VERSION : 0.1
   STRUCT
      SDC_Interlocks_In : "UDT_AB_Interlocks_SDC_In";
      SDC_Interlocks_Out : "UDT_AB_Interlocks_SDC_Out";
      Carrier : Array[1..99] of "UDT_AB_Interlocks_Carrier";
   END_STRUCT;
END_TYPE

TYPE "UDT_AB_Interlocks_SDC_Out"
VERSION : 0.1
   STRUCT
      SDC_Faulted : Bool;
      SDC_Status_1 : Bool;
      SDC_Status_2 : Bool;
      SDC_Status_3 : Bool;
      SDC_Status_4 : Bool;
      SDC_Status_5 : Bool;
      SDC_Status_6 : Bool;
      SDC_Status_7 : Bool;
      SDC_Status_8 : Bool;
      SDC_Status_9 : Bool;
      SDC_Status_10 : Bool;
      SDC_Status_11 : Bool;
      SDC_Status_12 : Bool;
      SDC_Status_13 : Bool;
      SDC_Status_14 : Bool;
      Heartbeat : Bool;
   END_STRUCT;
END_TYPE

// folder: UserDiag

TYPE "UserDiag_typeDevice"
TITLE = UserDiag_typeDevice
VERSION : 0.1
   STRUCT
      hardwareId : Hw_Device := 16#0000;   // Hardware identifier of the device/slave
      number : UInt := 0;   // Profinet device number/Profibus address of the slave
      "name" : String[50];   // Name of the device/slave
      ipAddress : IP_V4;   // IP address of the device
      state : USInt := 0;   // Status of the device/slave. 1:ok; 2:faulty, 3:lost connection, 4:disabled, 5:problem, 12:was faulty, 13:was lost, 14:was disabled, 15:problem gone
      exists : Bool := FALSE;   // TRUE: Device/slave is existing
      configured : Bool := FALSE;   // TRUE: Device/slave is configured
      faulty : Bool := FALSE;   // TRUE: Device/slave is faulty
      problem : Bool := FALSE;   // TRUE: Device/slave has a problem
      disabled : Bool := FALSE;   // TRUE: Device/slave is disabled
      error : Bool := FALSE;   // TRUE: Error in device/slave
      nextDevice : Int;   // device number of next device
      actualConfiguredSlots : Int := 0;   // Number of configured slots in the device/slave
      slots : Array[0.."USERDIAG_SLOTS_PER_DEVICE_UPPER_LIM"] of "UserDiag_typeSlot";   // Slot information of a device/slave
   END_STRUCT;
END_TYPE

TYPE "UserDiag_typeIOSystem"
TITLE = UserDiag_typeIOSystem
VERSION : 0.1
   STRUCT
      hardwareId : Hw_IoSystem := 16#0000;   // Hardware identifier of the IO-System/DP-Mastersystem
      number : UInt := 0;   // IO-System/DP-Mastersystem number
      error : Bool := FALSE;   // TRUE: Error in IO-System/DP-Mastersystem
      firstDevice : Int := 0;   // device number (index) of first device in IO System
      lastDevice : Int := 0;   // device number (index) of last device IO System
      actualConfiguredDevices : Int := 0;   // Number of configured devices/slaves in IO-System/DP-Mastersystem
      devices : Array[1.."USERDIAG_DEVICES_PER_IO_SYSTEM_UPPER_LIM"] of "UserDiag_typeDevice";   // Device/Slave information
   END_STRUCT;
END_TYPE

TYPE "UserDiag_typeActIOSystem"
TITLE = UserDiag_typeActIOSystem
VERSION : 0.1
   STRUCT
      actIOSystemNumber : Int := 1;   // Number of actual selected IO-system/DP-Mastersystem
      actIODeviceNumbers : Array[1.."USERDIAG_DEVICES_PER_SCREEN_UPPER_LIM"] of UInt;   // Device numbers/profibus addresses of actual selected IO-System/DP-Mastersystem
      actIODeviceState : Array[1.."USERDIAG_DEVICES_PER_SCREEN_UPPER_LIM"] of USInt;   // State of devices/slaves in actual selected IO-System/DP-Mastersystem
      actDeviceSlotsUsed : Array[0.."USERDIAG_SLOTS_PER_SCREEN_UPPER_LIM"] of Bool;   // Used slots of actual selected device/slave
      actDeviceSlotsState : Array[0.."USERDIAG_SLOTS_PER_SCREEN_UPPER_LIM"] of USInt;   // States of actual selected device/slave
   END_STRUCT;
END_TYPE

TYPE "UserDiag_typeHmiData"
VERSION : 0.1
   STRUCT
      actIOSystem : Int := 1;   // Index of actual selected IO-System/DP-Mastersystem
      actDeviceOfScreen : Int := 1;   // Index of selected device/slave on actual Screen
      ioSlotDiagnosticsLoaded : Bool;   // TRUE: Page for slot diagnostics is loaded
      actScreenDevices : Int := 1;   // Actual screennumber for copying device status to HMI
      maxScreensDevices : Int;   // Maximum screennumber for copying device status to HMI
      ackWaitTime : Int;   // Wait time after startup, for auto acknowledge
      ackStates : Bool;   // TRUE: Acknowledge of occurred errors in device/slave
      actIOSystemData : "UserDiag_typeActIOSystem";   // Data of actual IO system
      actDeviceNumber : UInt;   // Actual number/profibus address of device/slave
      actDeviceName : String[50];   // Name of actual selected device/slave
      actIPAddress : IP_V4;   // IP address of the device
      errorAtLowerScreen : Bool;   // Error at lower screen
      errorAtUpperScreen : Bool;   // Error at upper screen
      filterErrorDevices : Bool;   // Filter only fault devices
      ioSystemError : Array[1.."USERDIAG_IO_SYSTEMS_UPPER_LIM"] of Bool;   // Error in IO systems
   END_STRUCT;
END_TYPE

TYPE "UserDiag_typeSlot"
TITLE = UserDiag_typeSlot
VERSION : 0.1
   STRUCT
      hardwareId : Hw_Io := 16#0000;   // Hardware identifier of the module which is inserted in the slot
      state : USInt := 0;   // Status of the device/slave. 1:ok; 2:faulty, 3:lost connection, 4:disabled, 5:problem, 12:was faulty, 13:was lost, 14:was disabled, 15:problem gone
      exists : Bool := FALSE;   // TRUE: Modul is existing
      configured : Bool := FALSE;   // TRUE: Modul is configured
      faulty : Bool := FALSE;   // TRUE: Modul is faulty
      problem : Bool := FALSE;   // TRUE: Modul has a problem
      disabled : Bool := FALSE;   // TRUE: Modul is disabled
      error : Bool := FALSE;   // TRUE: Error in module which is inserted in the slot
   END_STRUCT;
END_TYPE

TYPE "UserDiag_typePLC"
TITLE = UserDiag_typePLC
VERSION : 0.1
   STRUCT
      hardwareId : Hw_Device := 16#0000;   // Hardware identifier of the PLC
      error : Bool := FALSE;   // TRUE: Error in PLC
      actualConfiguredSlots : Int := 0;   // Number of configured local slots at PLC
      slots : Array[0.."USERDIAG_SLOTS_PER_PLC_UPPER_LIM"] of "UserDiag_typeSlot";   // Information of the PLC slots; index = slotnumber; PLC always at slot 1
   END_STRUCT;
END_TYPE

// folder: 05_DBs

DATA_BLOCK "DB_SDC_TS_IF_COM_LOE"   // DB4
{ S7_Optimized_Access := 'FALSE' }
VERSION : 0.1
   VAR
      LoeSEK : "UDT_SDC_EMS_TS_COM";
   END_VAR
BEGIN
END_DATA_BLOCK

DATA_BLOCK "EMS"   // DB8
{ S7_Optimized_Access := 'TRUE' }
VERSION : 0.1
BEGIN
END_DATA_BLOCK

DATA_BLOCK "DB11_CARRIER"   // DB11
{ S7_Optimized_Access := 'TRUE' }
VERSION : 0.1
BEGIN
END_DATA_BLOCK

DATA_BLOCK "DB14_CarrZnFindArrayBuffer"   // DB14
{ S7_Optimized_Access := 'TRUE' }
VERSION : 0.1
BEGIN
END_DATA_BLOCK

DATA_BLOCK "DB15__FB_Zone_DB"   // DB15
{ S7_Optimized_Access := 'FALSE' }
VERSION : 0.1
"FB115_FB_Zone"
BEGIN
END_DATA_BLOCK

DATA_BLOCK "DB16_EMS_Status"   // DB16
{ S7_Optimized_Access := 'TRUE' }
VERSION : 0.1
   VAR
      EMS_DeviceStates : Struct
         Profinet1_Lddr : Hw_IoSystem := 257;
         DeviceStates_Mode2 : UInt := 2;
         DeviceStates_Mode4 : UInt := 4;
         DeviceStates_Mode5 : UInt := 5;
         DeviceStates_RetVal_2 : Int;
         DeviceStates_RetVal_4 : Int;
         DeviceStates_RetVal_5 : Int;
         DeviceStates_State2 : Array[0..1023] of Bool;
         DeviceStates_State4 : Array[0..1023] of Bool;
         DeviceStates_State5 : Array[0..1023] of Bool;
         DeviceStates_Condition_HMI : Array[0..82] of Int;
      END_STRUCT;
   END_VAR
BEGIN
END_DATA_BLOCK

DATA_BLOCK "TC_SDC_Out"   // DB53
{ S7_Optimized_Access := 'TRUE' }
VERSION : 0.1
BEGIN
END_DATA_BLOCK

DATA_BLOCK "DB101_DB_SDC_FAULTS"   // DB101
{ S7_Optimized_Access := 'FALSE' }
VERSION : 0.1
   VAR
      SDC_Fault : Word;
      Carrier_Fault : Array[1..90] of Word;
   END_VAR
BEGIN
END_DATA_BLOCK

DATA_BLOCK "DB110_DB_SDC_IN"   // DB110
{ S7_Optimized_Access := 'TRUE' }
VERSION : 0.1
   VAR
      Carrier : Array[0..99] of "UDT_SDC_IN";
   END_VAR
BEGIN
END_DATA_BLOCK

DATA_BLOCK "DB111_DB_SDC_OUT"   // DB111
{ S7_Optimized_Access := 'TRUE' }
VERSION : 0.1
   VAR
      Carrier : Array[0..99] of "UDT_SDC_OUT";
   END_VAR
BEGIN
END_DATA_BLOCK

DATA_BLOCK "DB116_TC_ZoneMotionControl"   // DB116
{ S7_Optimized_Access := 'TRUE' }
VERSION : 0.1
BEGIN
END_DATA_BLOCK

DATA_BLOCK "DB302_HMI_Faults"   // DB302
{ S7_Optimized_Access := 'TRUE' }
VERSION : 0.1
   VAR
      SDC_Faults_0 : Int := 0;
      SDC_Faults_1 : Int := 0;
      SDC_Faults_2 : Int := 0;
      SDC_Faults_3 : Int := 0;
      Carrier1_Faults_0 : Int := 0;
      Carrier1_Faults_1 : Int := 0;
      Carrier1_Faults_2 : Int := 0;
      Carrier1_Faults_3 : Int := 0;
      Carrier2_Faults_0 : Int := 0;
      Carrier2_Faults_1 : Int := 0;
      Carrier2_Faults_2 : Int := 0;
      Carrier2_Faults_3 : Int := 0;
      Carrier3_Faults_0 : Int := 0;
      Carrier3_Faults_1 : Int := 0;
      Carrier3_Faults_2 : Int := 0;
      Carrier3_Faults_3 : Int := 0;
      Carrier4_Faults_0 : Int := 0;
      Carrier4_Faults_1 : Int := 0;
      Carrier4_Faults_2 : Int := 0;
      Carrier4_Faults_3 : Int := 0;
      Carrier5_Faults_0 : Int := 1;
      Carrier5_Faults_1 : Int := 2;
      Carrier5_Faults_2 : Int := 3;
      Carrier5_Faults_3 : Int := 4;
      Carrier6_Faults_0 : Int := 5;
      Carrier6_Faults_1 : Int := 6;
      Carrier6_Faults_2 : Int := 7;
      Carrier6_Faults_3 : Int := 8;
      Carrier7_Faults_0 : Int := 9;
      Carrier7_Faults_1 : Int := 10;
      Carrier7_Faults_2 : Int := 11;
      Carrier7_Faults_3 : Int := 12;
      Carrier8_Faults_0 : Int := 13;
      Carrier8_Faults_1 : Int := 14;
      Carrier8_Faults_2 : Int := 15;
      Carrier8_Faults_3 : Int := 16;
      Carrier9_Faults_0 : Int := 17;
      Carrier9_Faults_1 : Int := 18;
      Carrier9_Faults_2 : Int := 19;
      Carrier9_Faults_3 : Int := 20;
      Carrier10_Faults_0 : Int := 21;
      Carrier10_Faults_1 : Int := 22;
      Carrier10_Faults_2 : Int := 23;
      Carrier10_Faults_3 : Int := 24;
      Carrier11_Faults_0 : Int := 25;
      Carrier11_Faults_1 : Int := 26;
      Carrier11_Faults_2 : Int := 27;
      Carrier11_Faults_3 : Int := 28;
      Carrier12_Faults_0 : Int := 29;
      Carrier12_Faults_1 : Int := 30;
      Carrier12_Faults_2 : Int := 31;
      Carrier12_Faults_3 : Int := 32;
      Carrier13_Faults_0 : Int := 33;
      Carrier13_Faults_1 : Int := 34;
      Carrier13_Faults_2 : Int := 35;
      Carrier13_Faults_3 : Int := 36;
      Carrier14_Faults_0 : Int := 37;
      Carrier14_Faults_1 : Int := 38;
      Carrier14_Faults_2 : Int := 39;
      Carrier14_Faults_3 : Int := 40;
      Carrier15_Faults_0 : Int := 41;
      Carrier15_Faults_1 : Int := 42;
      Carrier15_Faults_2 : Int := 43;
      Carrier15_Faults_3 : Int := 44;
      Carrier16_Faults_0 : Int := 45;
      Carrier16_Faults_1 : Int := 46;
      Carrier16_Faults_2 : Int := 47;
      Carrier16_Faults_3 : Int := 48;
      Carrier17_Faults_0 : Int := 49;
      Carrier17_Faults_1 : Int := 50;
      Carrier17_Faults_2 : Int := 51;
      Carrier17_Faults_3 : Int := 52;
      Carrier18_Faults_0 : Int := 53;
      Carrier18_Faults_1 : Int := 54;
      Carrier18_Faults_2 : Int := 55;
      Carrier18_Faults_3 : Int := 56;
      Carrier19_Faults_0 : Int := 57;
      Carrier19_Faults_1 : Int := 58;
      Carrier19_Faults_2 : Int := 59;
      Carrier19_Faults_3 : Int := 60;
      Carrier20_Faults_0 : Int := 61;
      Carrier20_Faults_1 : Int := 62;
      Carrier20_Faults_2 : Int := 63;
      Carrier20_Faults_3 : Int := 64;
      Carrier21_Faults_0 : Int := 65;
      Carrier21_Faults_1 : Int := 66;
      Carrier21_Faults_2 : Int := 67;
      Carrier21_Faults_3 : Int := 68;
      Carrier22_Faults_0 : Int := 69;
      Carrier22_Faults_1 : Int := 70;
      Carrier22_Faults_2 : Int := 71;
      Carrier22_Faults_3 : Int := 72;
      Carrier23_Faults_0 : Int := 73;
      Carrier23_Faults_1 : Int := 74;
      Carrier23_Faults_2 : Int := 75;
      Carrier23_Faults_3 : Int := 76;
      Carrier24_Faults_0 : Int := 77;
      Carrier24_Faults_1 : Int := 78;
      Carrier24_Faults_2 : Int := 79;
      Carrier24_Faults_3 : Int := 80;
      Carrier25_Faults_0 : Int := 81;
      Carrier25_Faults_1 : Int := 82;
      Carrier25_Faults_2 : Int := 83;
      Carrier25_Faults_3 : Int := 84;
      Carrier26_Faults_0 : Int := 85;
      Carrier26_Faults_1 : Int := 86;
      Carrier26_Faults_2 : Int := 87;
      Carrier26_Faults_3 : Int := 88;
      Carrier27_Faults_0 : Int := 89;
      Carrier27_Faults_1 : Int := 90;
      Carrier27_Faults_2 : Int := 91;
      Carrier27_Faults_3 : Int := 92;
      Carrier28_Faults_0 : Int := 93;
      Carrier28_Faults_1 : Int := 94;
      Carrier28_Faults_2 : Int := 95;
      Carrier28_Faults_3 : Int := 96;
      Carrier29_Faults_0 : Int := 97;
      Carrier29_Faults_1 : Int := 98;
      Carrier29_Faults_2 : Int := 99;
      Carrier29_Faults_3 : Int := 100;
      Carrier30_Faults_0 : Int := 101;
      Carrier30_Faults_1 : Int := 102;
      Carrier30_Faults_2 : Int := 103;
      Carrier30_Faults_3 : Int := 104;
      Carrier31_Faults_0 : Int := 105;
      Carrier31_Faults_1 : Int := 106;
      Carrier31_Faults_2 : Int := 107;
      Carrier31_Faults_3 : Int := 108;
      Carrier32_Faults_0 : Int := 109;
      Carrier32_Faults_1 : Int := 110;
      Carrier32_Faults_2 : Int := 111;
      Carrier32_Faults_3 : Int := 112;
      Carrier33_Faults_0 : Int := 113;
      Carrier33_Faults_1 : Int := 114;
      Carrier33_Faults_2 : Int := 115;
      Carrier33_Faults_3 : Int := 116;
      Carrier34_Faults_0 : Int := 117;
      Carrier34_Faults_1 : Int := 118;
      Carrier34_Faults_2 : Int := 119;
      Carrier34_Faults_3 : Int := 120;
      Carrier35_Faults_0 : Int := 121;
      Carrier35_Faults_1 : Int := 122;
      Carrier35_Faults_2 : Int := 123;
      Carrier35_Faults_3 : Int := 124;
      Carrier36_Faults_0 : Int := 125;
      Carrier36_Faults_1 : Int := 126;
      Carrier36_Faults_2 : Int := 127;
      Carrier36_Faults_3 : Int := 128;
      Carrier37_Faults_0 : Int := 129;
      Carrier37_Faults_1 : Int := 130;
      Carrier37_Faults_2 : Int := 131;
      Carrier37_Faults_3 : Int := 132;
      Carrier38_Faults_0 : Int := 133;
      Carrier38_Faults_1 : Int := 134;
      Carrier38_Faults_2 : Int := 135;
      Carrier38_Faults_3 : Int := 136;
      Carrier39_Faults_0 : Int := 137;
      Carrier39_Faults_1 : Int := 138;
      Carrier39_Faults_2 : Int := 139;
      Carrier39_Faults_3 : Int := 140;
      Carrier40_Faults_0 : Int := 141;
      Carrier40_Faults_1 : Int := 142;
      Carrier40_Faults_2 : Int := 143;
      Carrier40_Faults_3 : Int := 144;
      Carrier41_Faults_0 : Int := 145;
      Carrier41_Faults_1 : Int := 146;
      Carrier41_Faults_2 : Int := 147;
      Carrier41_Faults_3 : Int := 148;
      Carrier42_Faults_0 : Int := 149;
      Carrier42_Faults_1 : Int := 150;
      Carrier42_Faults_2 : Int := 151;
      Carrier42_Faults_3 : Int := 152;
      Carrier43_Faults_0 : Int := 153;
      Carrier43_Faults_1 : Int := 154;
      Carrier43_Faults_2 : Int := 155;
      Carrier43_Faults_3 : Int := 156;
      Carrier44_Faults_0 : Int := 157;
      Carrier44_Faults_1 : Int := 158;
      Carrier44_Faults_2 : Int := 159;
      Carrier44_Faults_3 : Int := 160;
      Carrier45_Faults_0 : Int := 161;
      Carrier45_Faults_1 : Int := 162;
      Carrier45_Faults_2 : Int := 163;
      Carrier45_Faults_3 : Int := 164;
      Carrier46_Faults_0 : Int := 165;
      Carrier46_Faults_1 : Int := 166;
      Carrier46_Faults_2 : Int := 167;
      Carrier46_Faults_3 : Int := 168;
      Carrier47_Faults_0 : Int := 169;
      Carrier47_Faults_1 : Int := 170;
      Carrier47_Faults_2 : Int := 171;
      Carrier47_Faults_3 : Int := 172;
      Carrier48_Faults_0 : Int := 173;
      Carrier48_Faults_1 : Int := 174;
      Carrier48_Faults_2 : Int := 175;
      Carrier48_Faults_3 : Int := 176;
      Carrier49_Faults_0 : Int := 177;
      Carrier49_Faults_1 : Int := 178;
      Carrier49_Faults_2 : Int := 179;
      Carrier49_Faults_3 : Int := 180;
      Carrier50_Faults_0 : Int := 181;
      Carrier50_Faults_1 : Int := 182;
      Carrier50_Faults_2 : Int := 183;
      Carrier50_Faults_3 : Int := 184;
      Carrier51_Faults_0 : Int := 185;
      Carrier51_Faults_1 : Int := 186;
      Carrier51_Faults_2 : Int := 187;
      Carrier51_Faults_3 : Int := 188;
      Carrier52_Faults_0 : Int := 189;
      Carrier52_Faults_1 : Int := 190;
      Carrier52_Faults_2 : Int := 191;
      Carrier52_Faults_3 : Int := 192;
      Carrier53_Faults_0 : Int := 193;
      Carrier53_Faults_1 : Int := 194;
      Carrier53_Faults_2 : Int := 195;
      Carrier53_Faults_3 : Int := 196;
      Carrier54_Faults_0 : Int := 197;
      Carrier54_Faults_1 : Int := 198;
      Carrier54_Faults_2 : Int := 199;
      Carrier54_Faults_3 : Int := 200;
      Carrier55_Faults_0 : Int := 201;
      Carrier55_Faults_1 : Int := 202;
      Carrier55_Faults_2 : Int := 203;
      Carrier55_Faults_3 : Int := 204;
      Carrier56_Faults_0 : Int := 205;
      Carrier56_Faults_1 : Int := 206;
      Carrier56_Faults_2 : Int := 207;
      Carrier56_Faults_3 : Int := 208;
      Carrier57_Faults_0 : Int := 209;
      Carrier57_Faults_1 : Int := 210;
      Carrier57_Faults_2 : Int := 211;
      Carrier57_Faults_3 : Int := 212;
      Carrier58_Faults_0 : Int := 213;
      Carrier58_Faults_1 : Int := 214;
      Carrier58_Faults_2 : Int := 215;
      Carrier58_Faults_3 : Int := 216;
      Carrier59_Faults_0 : Int := 217;
      Carrier59_Faults_1 : Int := 218;
      Carrier59_Faults_2 : Int := 219;
      Carrier59_Faults_3 : Int := 220;
      Carrier60_Faults_0 : Int := 221;
      Carrier60_Faults_1 : Int := 222;
      Carrier60_Faults_2 : Int := 223;
      Carrier60_Faults_3 : Int := 224;
      Carrier61_Faults_0 : Int := 225;
      Carrier61_Faults_1 : Int := 226;
      Carrier61_Faults_2 : Int := 227;
      Carrier61_Faults_3 : Int := 228;
      Carrier62_Faults_0 : Int := 229;
      Carrier62_Faults_1 : Int := 230;
      Carrier62_Faults_2 : Int := 231;
      Carrier62_Faults_3 : Int := 232;
      Carrier63_Faults_0 : Int := 233;
      Carrier63_Faults_1 : Int := 234;
      Carrier63_Faults_2 : Int := 235;
      Carrier63_Faults_3 : Int := 236;
      Carrier64_Faults_0 : Int := 237;
      Carrier64_Faults_1 : Int := 238;
      Carrier64_Faults_2 : Int := 239;
      Carrier64_Faults_3 : Int := 240;
      Carrier65_Faults_0 : Int := 241;
      Carrier65_Faults_1 : Int := 242;
      Carrier65_Faults_2 : Int := 243;
      Carrier65_Faults_3 : Int := 244;
      Carrier66_Faults_0 : Int := 245;
      Carrier66_Faults_1 : Int := 246;
      Carrier66_Faults_2 : Int := 247;
      Carrier66_Faults_3 : Int := 248;
      Carrier67_Faults_0 : Int := 249;
      Carrier67_Faults_1 : Int := 250;
      Carrier67_Faults_2 : Int := 251;
      Carrier67_Faults_3 : Int := 252;
      Carrier68_Faults_0 : Int := 253;
      Carrier68_Faults_1 : Int := 254;
      Carrier68_Faults_2 : Int := 255;
      Carrier68_Faults_3 : Int := 256;
      Carrier69_Faults_0 : Int := 257;
      Carrier69_Faults_1 : Int := 258;
      Carrier69_Faults_2 : Int := 259;
      Carrier69_Faults_3 : Int := 260;
      Carrier70_Faults_0 : Int := 261;
      Carrier70_Faults_1 : Int := 262;
      Carrier70_Faults_2 : Int := 263;
      Carrier70_Faults_3 : Int := 264;
      Carrier71_Faults_0 : Int := 265;
      Carrier71_Faults_1 : Int := 266;
      Carrier71_Faults_2 : Int := 267;
      Carrier71_Faults_3 : Int := 268;
      Carrier72_Faults_0 : Int := 269;
      Carrier72_Faults_1 : Int := 270;
      Carrier72_Faults_2 : Int := 271;
      Carrier72_Faults_3 : Int := 272;
      Carrier73_Faults_0 : Int := 273;
      Carrier73_Faults_1 : Int := 274;
      Carrier73_Faults_2 : Int := 275;
      Carrier73_Faults_3 : Int := 276;
      Carrier74_Faults_0 : Int := 277;
      Carrier74_Faults_1 : Int := 278;
      Carrier74_Faults_2 : Int := 279;
      Carrier74_Faults_3 : Int := 280;
      Carrier75_Faults_0 : Int := 281;
      Carrier75_Faults_1 : Int := 282;
      Carrier75_Faults_2 : Int := 283;
      Carrier75_Faults_3 : Int := 284;
      Carrier76_Faults_0 : Int := 285;
      Carrier76_Faults_1 : Int := 286;
      Carrier76_Faults_2 : Int := 287;
      Carrier76_Faults_3 : Int := 288;
      Carrier77_Faults_0 : Int := 289;
      Carrier77_Faults_1 : Int := 290;
      Carrier77_Faults_2 : Int := 291;
      Carrier77_Faults_3 : Int := 292;
      Carrier78_Faults_0 : Int := 293;
      Carrier78_Faults_1 : Int := 294;
      Carrier78_Faults_2 : Int := 295;
      Carrier78_Faults_3 : Int := 296;
      Carrier79_Faults_0 : Int := 297;
      Carrier79_Faults_1 : Int := 298;
      Carrier79_Faults_2 : Int := 299;
      Carrier79_Faults_3 : Int := 300;
      Carrier80_Faults_0 : Int := 301;
      Carrier80_Faults_1 : Int := 302;
      Carrier80_Faults_2 : Int := 303;
      Carrier80_Faults_3 : Int := 304;
      Carrier81_Faults_0 : Int := 305;
      Carrier81_Faults_1 : Int := 306;
      Carrier81_Faults_2 : Int := 307;
      Carrier81_Faults_3 : Int := 308;
      Carrier82_Faults_0 : Int := 309;
      Carrier82_Faults_1 : Int := 310;
      Carrier82_Faults_2 : Int := 311;
      Carrier82_Faults_3 : Int := 312;
   END_VAR
BEGIN
END_DATA_BLOCK

DATA_BLOCK "DB401_HMI_Status"   // DB401
{ S7_Optimized_Access := 'TRUE' }
VERSION : 0.1
   VAR
      Drive : "UDT_Drive_HMI";
      IO : "UDT_Carrier_IO_HMI";
      Status : "UDT_Carrier_Status_HMI";
      ZoneStatus : "UDT_Zone_Status_HMI";
   END_VAR
BEGIN
END_DATA_BLOCK

DATA_BLOCK "DB402_SDC_CARRIER_DRIVE_DATA"   // DB402
{ S7_Optimized_Access := 'TRUE' }
VERSION : 0.1
   VAR
      Drive_Data : "UDT_Carrier_Drive_Data";
   END_VAR
BEGIN
END_DATA_BLOCK

DATA_BLOCK "DB403_SDC_CARRIER_IO"   // DB403
{ S7_Optimized_Access := 'TRUE' }
VERSION : 0.1
   VAR
      IO_Data : "UDT_Carrier_IO_Data";
   END_VAR
BEGIN
END_DATA_BLOCK

DATA_BLOCK "Data_block_DO_NOT_CHANGE"   // DB999
{ S7_Optimized_Access := 'TRUE' }
VERSION : 0.1
   VAR RETAIN
      Production_Spacing_Memory : Int;
      Carrier_Spacing_Memory : Int;
   END_VAR
BEGIN
END_DATA_BLOCK

DATA_BLOCK "DB1000_AB_Interlocks"   // DB1000
{ S7_Optimized_Access := 'TRUE' }
VERSION : 0.1
   VAR
      Interlock : "UDT_AB_Interlocks";
   END_VAR
BEGIN
END_DATA_BLOCK

DATA_BLOCK "DB_SDC_GLOBAL"   // DB3700
{ S7_Optimized_Access := 'FALSE' }
AUTHOR : FFM
FAMILY : SDC
NAME : GLOBAL
VERSION : 1.0
   VAR
      EMS_ID_ACT : Int := 130;   // Aktuelle Anzahl der EMS-Treiber
      EMS_ID_MIN : Int := 1;   // Minimum EMS ID
      EMS_ID_MAX : Int := 184;   // Maximum EMS ID
      min_barcode_mm : DInt := 900;   // Lower limit, bar code value
      max_barcode_mm : DInt := 2076000;   // Upper limit, bar code value
      START_COURSE : DInt := 5800;   // Start Barcodevalue of Course
      END_COURSE : DInt := 312200;   // Ende Barcodewert vom Kurs
      SEK_MIN : Int := 1;   // Erste Abschnitt Nummer
      SEK_MAX : Int := 508;   // Aktuelle Anzahl der Bahnabschnitte
      TAKT_TIME : Int := 0;   // Reserve
      SEK_CYCLE_COUNTER : Int := 423;   // Section for increasing the track cycle counter
      MAN_V_1 : DInt := 6000;   // manual mode, set value: drive speed (mm/min)
      MAN_V_2 : DInt := 6000;   // manual mode, set value: drive speed (mm/min)
      min_Sequence_monitor_mm : DInt := 0;   // Lower limit of bar code value for sequence monitoring
      max_Sequence_monitor_mm : DInt := 0;   // Upper limit of bar code value for sequence monitoring
      MAX_PROFIL : Int := 10;   // maximal Profil Numbers
      CURR_EMS_ID_MAX : Int := 184;   // derzeit höchsten EMS-Nummer aktiv
      current_EMS_loop : Int := 0;   // Aktuelle Anzahl der EMS-Treiber auf Schleife
      EMS_ID_BUSY : Int := 0;   // EMS Driver wird aktiviert oder deaktiviert
      TAKT_TIME_LAST : Int := 0;   // Reserve
      Reserve_56 : Array[56..59] of Byte;
      SEK_REPAIR_1 : Int := 473;   // Section for repair, reset "send to repair 1" bit
      SEK_REPAIR_2 : Int := 0;   // Section for repair, reset "send to repair 2" bit
      SEK_DIAG_1 : Int := 0;   // Section diagnosticstation 1
      SEK_DIAG_2 : Int := 0;   // Section diagnosticstation 2
      SEK_DIAG_3 : Int := 0;   // Section diagnosticstation 2
      SEK_REP_1_START : Int := 470;
      SEK_REP_1_ENDE : Int := 472;
      SEK_REP_2_START : Int := 475;
      SEK_REP_2_ENDE : Int := 475;
      INFO_REP_1_DIAG_1 : Int := 0;   // Info for Function Rep 1 at Dignosticstation 1
      INFO_REP_2_DIAG_1 : Int := 0;   // Info for Function Rep 2 at Dignosticstation 1
      INFO_REP_1_DIAG_2 : Int := 0;   // Info for Function Rep 1 at Dignosticstation 2
      INFO_REP_2_DIAG_2 : Int := 0;   // Info for Function Rep 2 at Dignosticstation 2
      INFO_REP_1_DIAG_3 : Int := 0;   // Info for Function Rep 1 at Dignosticstation 2
      INFO_REP_2_DIAG_3 : Int := 0;   // Info for Function Rep 2 at Dignosticstation 2
      EMS_VCleaner_1 : Int := 0;   // EMS mit Vaccumreiniger No.1
      EMS_VCleaner_2 : Int := 0;   // EMS mit Vaccumreiniger No.2
      EMS_AKT_ZAEHLER_NR : Int := 131;   // EMS Aktualisierungsnummer
      EMS_AKT_ANZAHL : Int := 10;   // EMS Aktualisierunganzahl
      EMS_DIST_SEARCH : Int := 600;   // EMS Entfernungssuche zum vorderen EMS
      MIN_DIST_EMS : Array[0..15] of Int;   // minimum distance
      Reserve_132 : Array[132..149] of Byte;
      SYNCH : Array[0..15] of Struct   // Zur Abstandsregelung im Synchronbereich
         SET_DIST : Int;   // Set point value: distance (mm)
         SYNCH_DIST : Int;   // Start synchron distance value: distance (mm)
         HYST : Int;   // IO Hysterese
         K : Real;   // erreichen von Synchron Faktor
         MAX_FAKT : Real;   // Faktor für maximale Synchronisiergeschwindigkeit
         MIN_FAKT : Real;   // Faktor für minimale Synchronisiergeschwindigkeit
      END_STRUCT;
      Reserve_438 : Array[438..499] of Byte;   // spare
      LIMITS : Array[0..15] of Struct
         RAPID_SLOW : Int;   // Umstellung Begrenzung auf Abstand (mm), Einschränkung
         SLOW_SPEED_FAKT : Real;   // Faktor Geschwindigkeit für langsame Drehzahl
      END_STRUCT;
      Reserve_596 : Array[596..599] of Byte;   // spare
      "M" : Struct
         NEUSTART : Bool := FALSE;
         T_NEUSTART : Bool := FALSE;
         F_RESET : Bool := FALSE;
         "EMS_Read-Write" : Bool := FALSE;
         SDC_ER_Reset : Bool := FALSE;
      END_STRUCT;
   END_VAR
BEGIN
   MIN_DIST_EMS[0] := 6000;
   MIN_DIST_EMS[1] := 5970;
   MIN_DIST_EMS[2] := 6100;
   MIN_DIST_EMS[3] := 6000;
   MIN_DIST_EMS[4] := 6050;
   MIN_DIST_EMS[5] := 6100;
   MIN_DIST_EMS[6] := 6500;
   MIN_DIST_EMS[7] := 6500;
   MIN_DIST_EMS[8] := 6000;
   MIN_DIST_EMS[9] := 6250;
   MIN_DIST_EMS[10] := 6500;
   MIN_DIST_EMS[11] := 7000;
   MIN_DIST_EMS[12] := 7500;
   MIN_DIST_EMS[13] := 5950;
   MIN_DIST_EMS[14] := 5980;
   MIN_DIST_EMS[15] := 6500;
   SYNCH[0].SET_DIST := 6080;
   SYNCH[1].SET_DIST := 6030;
   SYNCH[2].SET_DIST := 6150;
   SYNCH[3].SET_DIST := 6080;
   SYNCH[4].SET_DIST := 6090;
   SYNCH[5].SET_DIST := 6400;
   SYNCH[6].SET_DIST := 6400;
   SYNCH[7].SET_DIST := 6400;
   SYNCH[8].SET_DIST := 6100;
   SYNCH[9].SET_DIST := 6300;
   SYNCH[10].SET_DIST := 6600;
   SYNCH[11].SET_DIST := 7100;
   SYNCH[12].SET_DIST := 7600;
   SYNCH[13].SET_DIST := 6510;
   SYNCH[14].SET_DIST := 6510;
   SYNCH[15].SET_DIST := 6510;
   SYNCH[0].SYNCH_DIST := 6400;
   SYNCH[1].SYNCH_DIST := 6450;
   SYNCH[2].SYNCH_DIST := 18000;
   SYNCH[3].SYNCH_DIST := 6200;
   SYNCH[4].SYNCH_DIST := 12000;
   SYNCH[5].SYNCH_DIST := 12000;
   SYNCH[6].SYNCH_DIST := 12000;
   SYNCH[7].SYNCH_DIST := 12000;
   SYNCH[8].SYNCH_DIST := 10000;
   SYNCH[9].SYNCH_DIST := 10000;
   SYNCH[10].SYNCH_DIST := 10000;
   SYNCH[11].SYNCH_DIST := 10000;
   SYNCH[12].SYNCH_DIST := 10000;
   SYNCH[13].SYNCH_DIST := 6800;
   SYNCH[14].SYNCH_DIST := 6800;
   SYNCH[15].SYNCH_DIST := 6800;
   SYNCH[0].HYST := 10;
   SYNCH[1].HYST := 4;
   SYNCH[2].HYST := 4;
   SYNCH[0].K := 1.0;
   SYNCH[1].K := 1.0;
   SYNCH[2].K := 1.0;
   SYNCH[3].K := 1.0;
   SYNCH[4].K := 1.3;
   SYNCH[5].K := 0.2;
   SYNCH[6].K := 0.2;
   SYNCH[7].K := 0.2;
   SYNCH[8].K := 1.0;
   SYNCH[9].K := 1.0;
   SYNCH[10].K := 1.0;
   SYNCH[11].K := 1.0;
   SYNCH[12].K := 1.0;
   SYNCH[13].K := 1.0;
   SYNCH[14].K := 1.0;
   SYNCH[15].K := 1.0;
   SYNCH[0].MAX_FAKT := 1.1;
   SYNCH[1].MAX_FAKT := 1.4;
   SYNCH[2].MAX_FAKT := 20.0;
   SYNCH[3].MAX_FAKT := 1.0;
   SYNCH[4].MAX_FAKT := 4.0;
   SYNCH[5].MAX_FAKT := 1.2;
   SYNCH[6].MAX_FAKT := 1.2;
   SYNCH[7].MAX_FAKT := 1.2;
   SYNCH[8].MAX_FAKT := 1.0;
   SYNCH[9].MAX_FAKT := 1.0;
   SYNCH[10].MAX_FAKT := 1.0;
   SYNCH[11].MAX_FAKT := 1.0;
   SYNCH[12].MAX_FAKT := 1.0;
   SYNCH[13].MAX_FAKT := 1.0;
   SYNCH[14].MAX_FAKT := 1.0;
   SYNCH[15].MAX_FAKT := 1.0;
   SYNCH[0].MIN_FAKT := 1.0;
   SYNCH[1].MIN_FAKT := 1.0;
   SYNCH[2].MIN_FAKT := 1.0;
   SYNCH[3].MIN_FAKT := 1.0;
   SYNCH[4].MIN_FAKT := 1.0;
   SYNCH[5].MIN_FAKT := 0.8;
   SYNCH[6].MIN_FAKT := 0.8;
   SYNCH[7].MIN_FAKT := 0.8;
   SYNCH[8].MIN_FAKT := 1.0;
   SYNCH[9].MIN_FAKT := 1.0;
   SYNCH[10].MIN_FAKT := 1.0;
   SYNCH[11].MIN_FAKT := 1.0;
   SYNCH[12].MIN_FAKT := 1.0;
   SYNCH[13].MIN_FAKT := 1.0;
   SYNCH[14].MIN_FAKT := 1.0;
   SYNCH[15].MIN_FAKT := 1.0;
   LIMITS[0].RAPID_SLOW := 7200;
   LIMITS[1].RAPID_SLOW := 7400;
   LIMITS[2].RAPID_SLOW := 7700;
   LIMITS[3].RAPID_SLOW := 8200;
   LIMITS[4].RAPID_SLOW := 8700;
   LIMITS[5].RAPID_SLOW := 6250;
   LIMITS[6].RAPID_SLOW := 7500;
   LIMITS[7].RAPID_SLOW := 7500;
   LIMITS[8].RAPID_SLOW := 6500;
   LIMITS[9].RAPID_SLOW := 6700;
   LIMITS[10].RAPID_SLOW := 7000;
   LIMITS[11].RAPID_SLOW := 7500;
   LIMITS[12].RAPID_SLOW := 8000;
   LIMITS[13].RAPID_SLOW := 6300;
   LIMITS[14].RAPID_SLOW := 6030;
   LIMITS[15].RAPID_SLOW := 7500;
   LIMITS[0].SLOW_SPEED_FAKT := 0.3;
   LIMITS[1].SLOW_SPEED_FAKT := 0.3;
   LIMITS[2].SLOW_SPEED_FAKT := 0.3;
   LIMITS[3].SLOW_SPEED_FAKT := 0.3;
   LIMITS[4].SLOW_SPEED_FAKT := 0.3;
   LIMITS[5].SLOW_SPEED_FAKT := 0.4;
   LIMITS[6].SLOW_SPEED_FAKT := 0.2;
   LIMITS[7].SLOW_SPEED_FAKT := 0.2;
   LIMITS[8].SLOW_SPEED_FAKT := 0.3;
   LIMITS[9].SLOW_SPEED_FAKT := 0.3;
   LIMITS[10].SLOW_SPEED_FAKT := 0.3;
   LIMITS[11].SLOW_SPEED_FAKT := 0.3;
   LIMITS[12].SLOW_SPEED_FAKT := 0.3;
   LIMITS[13].SLOW_SPEED_FAKT := 0.2;
   LIMITS[14].SLOW_SPEED_FAKT := 0.7;
   LIMITS[15].SLOW_SPEED_FAKT := 0.2;
   Reserve_132[132] := 16#00;
   Reserve_132[133] := 16#00;
   Reserve_132[134] := 16#00;
   Reserve_132[135] := 16#00;
   Reserve_132[136] := 16#00;
   Reserve_132[137] := 16#00;
   Reserve_132[138] := 16#00;
   Reserve_132[139] := 16#00;
   Reserve_132[140] := 16#00;
   Reserve_132[141] := 16#00;
   Reserve_132[142] := 16#00;
   Reserve_132[143] := 16#00;
   Reserve_132[144] := 16#00;
   Reserve_132[145] := 16#00;
   Reserve_132[146] := 16#00;
   Reserve_132[147] := 16#00;
   Reserve_132[148] := 16#00;
   Reserve_132[149] := 16#00;
   SYNCH[3].HYST := 4;
   SYNCH[4].HYST := 4;
   SYNCH[5].HYST := 0;
   SYNCH[6].HYST := 0;
   SYNCH[7].HYST := 0;
   SYNCH[8].HYST := 0;
   SYNCH[9].HYST := 0;
   SYNCH[10].HYST := 0;
   SYNCH[11].HYST := 0;
   SYNCH[12].HYST := 10;
   SYNCH[13].HYST := 4;
   SYNCH[14].HYST := 4;
   SYNCH[15].HYST := 4;
   Reserve_438[438] := 16#00;
   Reserve_438[439] := 16#00;
   Reserve_438[440] := 16#00;
   Reserve_438[441] := 16#00;
   Reserve_438[442] := 16#00;
   Reserve_438[443] := 16#00;
   Reserve_438[444] := 16#00;
   Reserve_438[445] := 16#00;
   Reserve_438[446] := 16#00;
   Reserve_438[447] := 16#00;
   Reserve_438[448] := 16#00;
   Reserve_438[449] := 16#00;
   Reserve_438[450] := 16#00;
   Reserve_438[451] := 16#00;
   Reserve_438[452] := 16#00;
   Reserve_438[453] := 16#00;
   Reserve_438[454] := 16#00;
   Reserve_438[455] := 16#00;
   Reserve_438[456] := 16#00;
   Reserve_438[457] := 16#00;
   Reserve_438[458] := 16#00;
   Reserve_438[459] := 16#00;
   Reserve_438[460] := 16#00;
   Reserve_438[461] := 16#00;
   Reserve_438[462] := 16#00;
   Reserve_438[463] := 16#00;
   Reserve_438[464] := 16#00;
   Reserve_438[465] := 16#00;
   Reserve_438[466] := 16#00;
   Reserve_438[467] := 16#00;
   Reserve_438[468] := 16#00;
   Reserve_438[469] := 16#00;
   Reserve_438[470] := 16#00;
   Reserve_438[471] := 16#00;
   Reserve_438[472] := 16#00;
   Reserve_438[473] := 16#00;
   Reserve_438[474] := 16#00;
   Reserve_438[475] := 16#00;
   // 32 more start values not shown
END_DATA_BLOCK

DATA_BLOCK "DB_SDC_EMS_FLAGS"   // DB3701
{ S7_Optimized_Access := 'FALSE' }
AUTHOR : FFM
FAMILY : SDC
NAME : GLOBAL